- PROFIenergy energy-saving mode active'; 8802 'A08802 - PROFIenergy not possible to switch off incremental encoder supply'; 13009 'F13009 - Licensing OA application not licensed'; 13100 'F13100 - Know-how protection: Copy protection error'; 13101 'F13101 - Know-how protection: Copy protection cannot be activated'; 13102 'F13102 - Know-how protection: Consistency error of the protected data'; 30001 'F30001 - Power unit: Overcurrent'; 30002 'F30002 - Power unit: DC link voltage overvoltage'; 30003 'F30003 - Power unit: DC link voltage undervoltage'; 30004 'F30004 - Power unit: Overtemperature heat sink AC inverter'; 30005 'F30005 - Power unit: Overload I2t'; 30011 'F30011 - Power unit: Line phase failure in main circuit'; 30015 'F30015 (N, A) - Power unit: Phase failure motor cable'; 30016 'A30016 (N) - Power unit: Load supply switched out'; 30017 'F30017 - Power unit: Hardware current limit has responded too often'; 30021 'F30021 - Power unit: Ground fault'; 30022 'F30022 - Power unit: Monitoring U_ce'; 30024 'F30024 - Power unit: Overtemperature thermal model'; 30025 'F30025 - Power unit: Chip overtemperature'; 30027 'F30027 - Power unit: Precharging DC link time monitoring'; 30031 'A30031 - Power unit: Hardware current limiting in phase U'; 30032 'A30032 - Power unit: Hardware current limiting in phase V'; 30033 'A30033 - Power unit: Hardware current limiting in phase W'; 30034 'A30034 - Power unit: Internal overtemperature'; 30042 'A30042 - Power unit: Fan has reached the maximum operating hours'; 30051 'F30051 - Power unit: Motor holding brake short circuit detected'; 30052 'F30052 - EEPROM data error'; 30054 'A30054 (F, N) - Power unit: Undervoltage when opening the brake'; 30057 'A30057 - Power unit: Line asymmetry'; 30065 'A30065 (F, N) - Voltage measured values not plausible'; 30071 'F30071 - No new actual values received from the Power Module'; 30072 'F30072 - Setpoints can no longer be transferred to the Power Module'; 30074 'F30074 (A) - Communication error between the Control Unit and Power Module'; 30075 'F30075 - Configuration of the power unit unsuccessful'; 30080 'F30080 - Power unit: Current increasing too quickly'; 30081 'F30081 - Power unit: Switching operations too frequent'; 30105 'F30105 - PU: Actual value sensing fault'; 30502 'A30502 - Power unit: DC link overvoltage'; 30600 'F30600 - SI P2: STOP A initiated'; 30611 'F30611 (A) - SI P2: Defect in a monitoring channel'; 30620 'N30620 (F, A) - SI P2: Safe Torque Off active'; 30625 'F30625 - SI P2: Sign-of-life error in safety data'; 30649 'F30649 - SI P2: Internal software error'; 30650 'F30650 - SI P2: Acceptance test required'; 30651 'F30651 - SI P2: Synchronization with Control Unit unsuccessful'; 30655 'F30655 - SI P2: Align monitoring functions'; 30656 'F30656 - SI P2: Parameter processor 2 parameter error'; 30659 'F30659 - SI P2: Write request for parameter rejected'; 30662 'F30662 - Error in internal communications'; 30664 'F30664 - Error while booting'; 30665 'F30665 - SI P2: System is defective'; 30666 'A30666 (F) - SI Motion P2: Steady-state (static) 1 signal at the F-DI for safe acknowledgment'; 30680 'F30680 - SI Motion P2: Checksum error safety monitoring functions'; 30681 'F30681 - SI Motion P1: Incorrect parameter value'; 30682 'F30682 - SI Motion P2: Monitoring function not supported'; 30683 'F30683 - SI Motion P2: SLS enable missing'; 30692 'F30692 - SI Motion P2: Parameter value not permitted for encoderless'; 30693 'A30693 (F) - SI P2: Safety parameter settings changed, POWER ON required'; 30700 'C30700 - SI Motion P2: STOP A initiated'; 30701 'C30701 - SI Motion P2: STOP B initiated'; 30706 'C30706 - SI Motion P2: SAM/SBR limit exceeded'; 30711 'C30711 - SI Motion P2: Defect in a monitoring channel'; 30712 'C30712 - SI Motion P2: Defect in F-IO processing'; 30714 'C30714 - SI Motion P2: Safely limited speed exceeded'; 30716 'C30716 - SI Motion P2: Tolerance for safe motion direction exceeded'; 30770 'C30770 - SI Motion P2: Discrepancy error affecting the failsafe inputs'; 30772 'A30772 - SI Motion P2: Test stop for fail-safe digital outputs running'; 30773 'F30773 - SI Motion P2: Test stop fail-safe digital output error'; 30788 'A30788 - Automatic test stop: wait for STO deselection via SMM'; 30798 'C30798 - SI Motion P2: Test stop for motion monitoring functions running'; 30799 'C30799 - SI Motion P2: Acceptance test mode active'; 30800 'N30800 (F) - Power unit: Group signal'; 30802 'F30802 - Power unit: Time slice overflow'; 30804 'F30804 (N, A) - Power unit: CRC'; 30805 'F30805 - Power unit: EEPROM checksum error'; 30809 'F30809 - Power unit: Switching information not valid'; 30810 'A30810 (F) - Power unit: Watchdog timer'; 30850 'F30850 - Power unit: Internal software error'; 30903 'F30903 - Power unit: I2C bus error occurred'; 30920 'A30920 (F) - Temperature sensor fault'; 30950 'F30950 - Power unit: Internal software error'; 30999 'A30999 (F, N) - Power unit: Unknown alarm'; 31100 'F31100 (N, A) - Encoder 1: Zero mark distance error'; 31101 'F31101 (N, A) - Encoder 1: Zero mark failed'; 31103 'F31103 (N, A) - Encoder 1: Amplitude error track R'; 31118 'F31118 (N, A) - Encoder 1: Speed difference outside the tolerance range'; 31131 'F31131 (N, A) - Encoder 1: Deviation position incremental/absolute too large'; 31150 'F31150 (N, A) - Encoder 1: Initialization error'; 31153 'F31153 (N, A) - Encoder 1: Identification error'; 31400 'A31400 (F, N) - Encoder 1: Alarm threshold zero mark distance error'; 31401 'A31401 (F, N) - Encoder 1: Alarm threshold zero mark failed'; 31418 'A31418 (F, N) - Encoder 1: Speed difference per sampling rate exceeded'; 31422 'A31422 (F, N) - Encoder 1: Pulses per revolution square-wave encoder outside tolerance bandwidth'; 31431 'A31431 (F, N) - Encoder 1: Deviation position incremental/absolute too large'; 31802 'F31802 (N, A) - Encoder 1: Time slice overflow'; 31805 'F31805 (N, A) - Encoder 1: EEPROM checksum error'; 31850 'F31850 (N, A) - Encoder 1: Encoder evaluation internal software error'; 31899 'F31899 (N, A) - Encoder 1: Unknown fault'; 31905 'F31905 (N, A) - Encoder 1: Parameterization error'; 31915 'A31915 (F, N) - Encoder 1: Configuration error'; 31930 'A31930 (N) - Encoder 1: Data logger has saved data'; 31950 'F31950 - Encoder 1: Internal software error'; 31999 'A31999 (F, N) - Encoder 1: Unknown alarm'; 32110 'F32110 (N, A) - Encoder 2: Serial communications error'; 32111 'F32111 (N, A) - Encoder 2: Absolute encoder internal fault'; 32112 'F32112 (N, A) - Encoder 2: Error bit set in the serial protocol'; 32150 'F32150 (N, A) - Encoder 2: Initialization error'; 32153 'F32153 (N, A) - Encoder 2: Identification error'; 32410 'A32410 (F, N) - Encoder 2: Serial communications'; 32411 'A32411 (F, N) - Encoder 2: Absolute encoder signals internal alarms'; 32412 'A32412 (F, N) - Encoder 2: Error bit set in the serial protocol'; 32442 'A32442 (F, N) - Encoder 2: Battery voltage pre-alarm'; 32802 'F32802 (N, A) - Encoder 2: Time slice overflow'; 32805 'F32805 (N, A) - Encoder 2: EEPROM checksum error'; 32850 'F32850 (N, A) - Encoder 2: Encoder evaluation internal software error'; 32899 'F32899 (N, A) - Encoder 2: Unknown fault'; 32905 'F32905 (N, A) - Encoder 2: Parameterization error'; 32915 'A32915 (F, N) - Encoder 2: Configuration error'; 32930 'A32930 (N) - Encoder 2: Data logger has saved data'; 32950 'F32950 - Encoder 2: Internal software error'; 32999 'A32999 (F, N) - Encoder 2: Unknown alarm'; 50001 'A50001 (F) - PROFINET configuration error'; 50010 'A50010 (F) - PROFINET: Consistency error affecting adjustable parameters'; 50011 'A50011 (F) - Ethernet/IP: configuration error'; 50020 'A50020 (F) - PROFINET: Second controller missing'; 50510 'F50510 - FBLOCKS: Logon of the run-time group rejected'; 50511 'F50511 - FBLOCKS: Memory no longer available for free function blocks'; 50513 'A50513 (F) - FBLOCKS: Run sequence value already assigned'; 50517 'A50517 - FBLOCKS: Int. meas. active'; 50518 'F50518 - FBLOCKS: Sampling time of free run-time group differs at download'

text list "SDC_FAULTS-Old": 11 'Carrier 1 PLC Not Communicating'; 12 'Carrier 2 PLC Not Communicating'; 13 'Carrier 3 PLC Not Communicating'; 14 'Carrier 4 PLC Not Communicating'; 21 'Carrier 1 Safe Input Card Fault'; 22 'Carrier 1 Safe Output Card Fault'; 23 'Carrier 1 Standard Input Card Fault'; 24 'Carrier 1 Standard Output Card Fault'; 25 'Carrier 2 Safe Input Card Fault'; 26 'Carrier 2 Safe Output Card Fault'; 27 'Carrier 2 Standard Input Card Fault'; 28 'Carrier 2 Standard Output Card Fault'; 29 'Carrier 3 Safe Input Card Fault'; 30 'Carrier 3 Safe Output Card Fault'; 31 'Carrier 3 Standard Input Card Fault'; 32 'Carrier 3 Standard Output Card Fault'; 33 'Carrier 4 Safe Input Card Fault'; 34 'Carrier 4 Safe Output Card Fault'; 35 'Carrier 4 Standard Input Card Fault'; 36 'Carrier 4 Standard Output Card Fault'; 51 'Carrier 1 VFD Drive Fault'; 52 'Carrier 2 VFD Drive Fault'; 53 'Carrier 3 VFD Drive Fault'; 54 'Carrier 4 VFD Drive Fault'; 502 'Carrier 2 Crash Detection Fault'; 201 'Carrier 1 Encoder Reader Tilted 180 Degrees'; 202 'Carrier 1 Encoder Position Error'; 203 'Carrier 1 Encoder Internal Fault'; 211 'Carrier 2 Encoder Reader Tilted 180 Degrees'; 212 'Carrier 2 Encoder Position Error'; 213 'Carrier 2 Encoder Internal Fault'; 221 'Carrier 3 Encoder Reader Tilted 180 Degrees'; 222 'Carrier 3 Encoder Position Error'; 223 'Carrier 3 Encoder Internal Fault'; 231 'Carrier 4 Encoder Reader Tilted 180 Degrees'; 232 'Carrier 4 Encoder Position Error'; 233 'Carrier 4 Encoder Internal Fault'; 101 'Carrier 1 CB2120 Tripped'; 102 'Carrier 1 CB2121 Tripped'; 103 'Carrier 1 CB2122 Tripped'; 104 'Carrier 1 CB2123 Tripped'; 131 'Carrier 4 CB2120 Tripped'; 132 'Carrier 4 CB2121 Tripped'; 133 'Carrier 4 CB2122 Tripped'; 134 'Carrier 4 CB2123 Tripped'; 111 'Carrier 2 CB2120 Tripped'; 112 'Carrier 2 CB2121 Tripped'; 113 'Carrier 2 CB2122 Tripped'; 114 'Carrier 2 CB2123 Tripped'; 121 'Carrier 3 CB2120 Tripped'; 122 'Carrier 3 CB2121 Tripped'; 123 'Carrier 3 CB2122 Tripped'; 124 'Carrier 3 CB2123 Tripped'

text list "SDC_FAULTS": 24 'Scalance Ethernet SW2 Comm Fault'; 100 'Carrier 1 Profinet Comms Fault'; 101 'Carrier 1 Disconnect Open Power Fault DI11.0'; 102 'Carrier 1 CB02120 Tripped'; 103 'Carrier 1 CB02121 Tripped'; 104 'Carrier 1 CB02122 Tripped'; 105 'Carrier 1 CB02123 Tripped'; 106 'Carrier 1 AUX1 CB Tripped DI11.4'; 107 'Carrier 1 AUX2 CB Tripped DI11.5'; 111 'Carrier 1 PLC Not Communicating'; 121 'Carrier 1 Safe Input Card Fault'; 122 'Carrier 1 Safe Output Card Fault'; 123 'Carrier 1 Standard Input Card Fault'; 124 'Carrier 1 Standard Output Card Fault'; 130 'Carrier 1 PF Reader Tilted 180°'; 131 'Carrier 1 PF Reader Internal Error'; 132 'Carrier 1 PF Reader Position Error'; 133 'Carrier 1 PF Reader Comm Fault'; 134 'Carrier 1 FR HMI Comm Fault'; 140 'Carrier 1 Crash Detection Fault'; 145 'Carrier 1 Carrier Number Invalid'; 150 'F01653 - Carrier 1 SI P1 (CU): PROFIBUS/PROFINET configuration error'; 151 'F01662 - Carrier 1 Error internal communications'; 160 'F07011 - Carrier 1 Drive: Motor overtemperature'; 161 'F07016 - Carrier 1 Drive: Motor temperature sensor fault'; 162 'F07801 - Carrier 1 Drive: Motor overcurrent'; 163 'F07802 - Carrier 1 Drive: Infeed or power unit not ready'; 164 'F07807 - Carrier 1 Drive: Short-circuit/ground fault detected'; 170 'F08501 - Carrier 1 PROFINET: Setpoint timeout'; 180 'F30001 - Carrier 1 Power unit: Overcurrent'; 181 'F30002 - Carrier 1 Power unit: DC link voltage overvoltage'; 182 'F30003 - Carrier 1 Power unit: DC link voltage undervoltage'; 183 'F30004 - Carrier 1 Power unit: Overtemperature heat sink AC inverter'; 184 'F30005 - Carrier 1 Power unit: Overload I2t'; 185 'F30011 - Carrier 1 Power unit: Line phase failure in main circuit'; 186 'F30015 - Carrier 1 Power unit: Phase failure motor cable'; 20 'Rockwell PLC Comm Fault'; 21 'WLAN1 Comm Fault'; 22 'WLAN2 Comm Fault'; 23 'Scalance Ethernet SW1 Comm Fault'; 187 'F30021 - Carrier 1 Power unit: Ground fault'; 188 'F30024 - Carrier 1 Power unit: Overtemperature thermal model'; 189 'F30051 - Carrier 1 Power unit: Motor holding brake short circuit detected'; 200 'Carrier 2 Profinet Comms Fault'; 201 'Carrier 2 Disconnect Open Power Fault DI11.0'; 202 'Carrier 2 CB02120 Tripped'; 203 'Carrier 2 CB02121 Tripped'; 204 'Carrier 2 CB02122 Tripped'; 205 'Carrier 2 CB02123 Tripped'; 206 'Carrier 2 AUX1 CB Tripped DI11.4'; 207 'Carrier 2 AUX2 CB Tripped DI11.5'; 211 'Carrier 2 PLC Not Communicating'; 221 'Carrier 2 Safe Input Card Fault'; 222 'Carrier 2 Safe Output Card Fault'; 223 'Carrier 2 Standard Input Card Fault'; 224 'Carrier 2 Standard Output Card Fault'; 230 'Carrier 2 PF Reader Tilted 180°'; 231 'Carrier 2 PF Reader Position Error'; 232 'Carrier 2 PF Reader Internal Error'; 233 'Carrier 2 PF Reader Comm Fault'; 234 'Carrier 2 FR HMI Comm Fault'; 240 'Carrier 2 Crash Detection Fault'; 245 'Carrier 2 Carrier Number Invalid'; 250 'F01653 - Carrier 2 SI P1 (CU): PROFIBUS/PROFINET configuration error'; 251 'F01662 - Carrier 2 Error internal communications'; 260 'F07011 - Carrier 2 Drive: Motor overtemperature'; 261 'F07016 - Carrier 2 Drive: Motor temperature sensor fault'; 262 'F07801 - Carrier 2 Drive: Motor overcurrent'; 263 'F07802 - Carrier 2 Drive: Infeed or power unit not ready'; 264 'F07807 - Carrier 2 Drive: Short-circuit/ground fault detected'; 270 'F08501 - Carrier 2 PROFINET: Setpoint timeout'; 280 'F30001 - Carrier 2 Power unit: Overcurrent'; 281 'F30002 - Carrier 2 Power unit: DC link voltage overvoltage'; 282 'F30003 - Carrier 2 Power unit: DC link voltage undervoltage'; 283 'F30004 - Carrier 2 Power unit: Overtemperature heat sink AC inverter'; 284 'F30005 - Carrier 2 Power unit: Overload I2t'; 285 'F30011 - Carrier 2 Power unit: Line phase failure in main circuit'; 286 'F30015 - Carrier 2 Power unit: Phase failure motor cable'; 287 'F30021 - Carrier 2 Power unit: Ground fault'; 288 'F30024 - Carrier 2 Power unit: Overtemperature thermal model'; 289 'F30051 - Carrier 2 Power unit: Motor holding brake short circuit detected'; 300 'Carrier 3 Profinet Comms Fault'; 301 'Carrier 3 Disconnect Open Power Fault DI11.0'; 302 'Carrier 3 CB02120 Tripped'; 303 'Carrier 3 CB02121 Tripped'; 304 'Carrier 3 CB02122 Tripped'; 305 'Carrier 3 CB02123 Tripped'; 306 'Carrier 3 AUX1 CB Tripped DI11.4'; 307 'Carrier 3 AUX2 CB Tripped DI11.5'; 311 'Carrier 3 PLC Not Communicating'; 321 'Carrier 3 Safe Input Card Fault'; 322 'Carrier 3 Safe Output Card Fault'; 323 'Carrier 3 Standard Input Card Fault'; 324 'Carrier 3 Standard Output Card Fault'; 330 'Carrier 3 PF Reader Tilted 180°'; 331 'Carrier 3 PF Reader Position Error'; 332 'Carrier 3 PF Reader Internal Error'; 333 'Carrier 3 PF Reader Comm Fault'; 334 'Carrier 3 FR HMI Comm Fault'; 340 'Carrier 3 Crash Detection Fault'; 345 'Carrier 3 Carrier Number Invalid'; 350 'F01653 - Carrier 3 SI P1 (CU): PROFIBUS/PROFINET configuration error'; 351 'F01662 - Carrier 3 Error internal communications'; 360 'F07011 - Carrier 3 Drive: Motor overtemperature'; 361 'F07016 - Carrier 3 Drive: Motor temperature sensor fault'; 362 'F07801 - Carrier 3 Drive: Motor overcurrent'; 363 'F07802 - Carrier 3 Drive: Infeed or power unit not ready'; 364 'F07807 - Carrier 3 Drive: Short-circuit/ground fault detected'; 370 'F08501 - Carrier 3 PROFINET: Setpoint timeout'; 380 'F30001 - Carrier 3 Power unit: Overcurrent'; 381 'F30002 - Carrier 3 Power unit: DC link voltage overvoltage'; 382 'F30003 - Carrier 3 Power unit: DC link voltage undervoltage'; 383 'F30004 - Carrier 3 Power unit: Overtemperature heat sink AC inverter'; 384 'F30005 - Carrier 3 Power unit: Overload I2t'; 385 'F30011 - Carrier 3 Power unit: Line phase failure in main circuit'; 386 'F30015 - Carrier 3 Power unit: Phase failure motor cable'; 387 'F30021 - Carrier 3 Power unit: Ground fault'; 388 'F30024 - Carrier 3 Power unit: Overtemperature thermal model'; 389 'F30051 - Carrier 3 Power unit: Motor holding brake short circuit detected'; 400 'Carrier 4 Profinet Comms Fault'; 401 'Carrier 4 Disconnect Open Power Fault DI11.0'; 402 'Carrier 4 CB02120 Tripped'; 403 'Carrier 4 CB02121 Tripped'; 404 'Carrier 4 CB02122 Tripped'; 405 'Carrier 4 CB02123 Tripped'; 406 'Carrier 4 AUX1 CB Tripped DI11.4'; 407 'Carrier 4 AUX2 CB Tripped DI11.5'; 411 'Carrier 4 PLC Not Communicating'; 421 'Carrier 4 Safe Input Card Fault'; 422 'Carrier 4 Safe Output Card Fault'; 423 'Carrier 4 Standard Input Card Fault'; 424 'Carrier 4 Standard Output Card Fault'; 430 'Carrier 4 PF Reader Tilted 180°'; 431 'Carrier 4 PF Reader Position Error'; 432 'Carrier 4 PF Reader Internal Error'; 433 'Carrier 4 PF Reader Comm Fault'; 434 'Carrier 4 FR HMI Comm Fault'; 440 'Carrier 4 Crash Detection Fault'; 445 'Carrier 4 Carrier Number Invalid'; 450 'F01653 - Carrier 4 SI P1 (CU): PROFIBUS/PROFINET configuration error'; 451 'F01662 - Carrier 4 Error internal communications'; 460 'F07011 - Carrier 4 Drive: Motor overtemperature'; 461 'F07016 - Carrier 4 Drive: Motor temperature sensor fault'; 462 'F07801 - Carrier 4 Drive: Motor overcurrent'; 463 'F07802 - Carrier 4 Drive: Infeed or power unit not ready'; 464 'F07807 - Carrier 4 Drive: Short-circuit/ground fault detected'; 470 'F08501 - Carrier 4 PROFINET: Setpoint timeout'; 480 'F30001 - Carrier 4 Power unit: Overcurrent'; 481 'F30002 - Carrier 4 Power unit: DC link voltage overvoltage'; 482 'F30003 - Carrier 4 Power unit: DC link voltage undervoltage'; 483 'F30004 - Carrier 4 Power unit: Overtemperature heat sink AC inverter'; 484 'F30005 - Carrier 4 Power unit: Overload I2t'; 485 'F30011 - Carrier 4 Power unit: Line phase failure in main circuit'; 486 'F30015 - Carrier 4 Power unit: Phase failure motor cable'; 487 'F30021 - Carrier 4 Power unit: Ground fault'; 488 'F30024 - Carrier 4 Power unit: Overtemperature thermal model'; 489 'F30051 - Carrier 4 Power unit: Motor holding brake short circuit detected'; 10 'Carrier Spacing Fault'

graphic list "Grafikliste_G_Y": 0 'Green pilot light 2'; 1 'Yellow pilot light 2'

graphic list "PB_Slave_Bit12_3": 0 'PB_Array_blau_3'; 1 'PB_Array_grün_3'

graphic list "PB_Slave_Bit10_3": 0 'PB_Array_blau_3'; 1 'PB_Array_grün_3'

graphic list "PB_Slave_Bit7_3": 0 'PB_Array_blau_3'; 1 'PB_Array_grün_3'

graphic list "PB_Slave_Bit6_3": 1 'PB_Array_grün_3'; 0 'PB_Array_blau_3'

graphic list "PB_Slave_Bit5_3": 0 'PB_Array_blau_3'; 1 'PB_Array_grün_3'

graphic list "PB_Slave_Bit1_3": 1 'PB_Array_grün_3'; 0 'PB_Array_blau_3'

graphic list "PB_Slave_Bit3_3": 1 'PB_Array_grün_3'; 0 'PB_Array_blau_3'

graphic list "PB_Slave_Bit9_3": 0 'PB_Array_blau_3'; 1 'PB_Array_grün_3'

graphic list "PB_Slave_Bit8_3": 1 'PB_Array_grün_3'; 0 'PB_Array_blau_3'

graphic list "PB_Slave_Bit0_3": 1 'PB_Array_grün_3'; 0 'PB_Array_blau_3'

graphic list "PB_Slave_Bit4_3": 1 'PB_Array_grün_3'; 0 'PB_Array_blau_3'

graphic list "PB_Slave_Bit14_3": 0 'PB_Array_blau_3'; 1 'PB_Array_grün_3'

graphic list "PB_Slave_Bit11_3": 0 'PB_Array_blau_3'; 1 'PB_Array_grün_3'

graphic list "PB_Slave_Bit2_3": 1 'PB_Array_grün_3'; 0 'PB_Array_blau_3'

graphic list "PB_Slave_Bit13_3": 0 'PB_Array_blau_3'; 1 'PB_Array_grün_3'

graphic list "PB_Slave_Bit15_3": 1 'PB_Array_grün_3'; 0 'PB_Array_blau_3'

graphic list "PB_Slave_Bit1_1": 1 'PB_Array_grün_1'; 0 'PB_Array_blau_1'

graphic list "PB_Slave_Bit0_1": 1 'PB_Array_grün_1'; 0 'PB_Array_blau_1'

graphic list "PB_Slave_Bit2_1": 1 'PB_Array_grün_1'; 0 'PB_Array_blau_1'

graphic list "PB_Slave_Bit4_1": 1 'PB_Array_grün_1'; 0 'PB_Array_blau_1'

graphic list "PB_Slave_Bit3_1": 1 'PB_Array_grün_1'; 0 'PB_Array_blau_1'

graphic list "PB_Slave_Bit5_1": 0 'PB_Array_blau_1'; 1 'PB_Array_grün_1'

graphic list "PB_Slave_Bit7_1": 0 'PB_Array_blau_1'; 1 'PB_Array_grün_1'

graphic list "PB_Slave_Bit6_1": 1 'PB_Array_grün_1'; 0 'PB_Array_blau_1'

graphic list "PB_Slave_Bit13_1": 0 'PB_Array_blau_1'; 1 'PB_Array_grün_1'

graphic list "PB_Slave_Bit10_1": 0 'PB_Array_blau_1'; 1 'PB_Array_grün_1'

graphic list "PB_Slave_Bit12_1": 0 'PB_Array_blau_1'; 1 'PB_Array_grün_1'

graphic list "PB_Slave_Bit15_1": 1 'PB_Array_grün_1'; 0 'PB_Array_blau_1'

graphic list "PB_Slave_Bit9_1": 0 'PB_Array_blau_1'; 1 'PB_Array_grün_1'

graphic list "PB_Slave_Bit8_1": 1 'PB_Array_grün_1'; 0 'PB_Array_blau_1'

graphic list "PB_Slave_Bit11_1": 0 'PB_Array_blau_1'; 1 'PB_Array_grün_1'

graphic list "PB_Slave_Bit14_1": 0 'PB_Array_blau_1'; 1 'PB_Array_grün_1'

graphic list "PB_Slave_Bit4_2": 1 'PB_Array_grün_2'; 0 'PB_Array_blau_2'

graphic list "PB_Slave_Bit5_2": 0 'PB_Array_blau_2'; 1 'PB_Array_grün_2'

graphic list "PB_Slave_Bit7_2": 0 'PB_Array_blau_2'; 1 'PB_Array_grün_2'

graphic list "PB_Slave_Bit6_2": 1 'PB_Array_grün_2'; 0 'PB_Array_blau_2'

graphic list "PB_Slave_Bit2_2": 1 'PB_Array_grün_2'; 0 'PB_Array_blau_2'

graphic list "PB_Slave_Bit3_2": 1 'PB_Array_grün_2'; 0 'PB_Array_blau_2'

graphic list "PB_Slave_Bit1_2": 1 'PB_Array_grün_2'; 0 'PB_Array_blau_2'

graphic list "PB_Slave_Bit0_2": 1 'PB_Array_grün_2'; 0 'PB_Array_blau_2'

graphic list "PB_Slave_Bit14_2": 0 'PB_Array_blau_2'; 1 'PB_Array_grün_2'

graphic list "PB_Slave_Bit12_2": 0 'PB_Array_blau_2'; 1 'PB_Array_grün_2'

graphic list "PB_Slave_Bit15_2": 1 'PB_Array_grün_2'; 0 'PB_Array_blau_2'

graphic list "PB_Slave_Bit13_2": 0 'PB_Array_blau_2'; 1 'PB_Array_grün_2'

graphic list "PB_Slave_Bit10_2": 0 'PB_Array_blau_2'; 1 'PB_Array_grün_2'

graphic list "PB_Slave_Bit9_2": 0 'PB_Array_blau_2'; 1 'PB_Array_grün_2'

graphic list "PB_Slave_Bit8_2": 1 'PB_Array_grün_2'; 0 'PB_Array_blau_2'

graphic list "PB_Slave_Bit11_2": 0 'PB_Array_blau_2'; 1 'PB_Array_grün_2'

graphic list "@DiagnosticsStates": 0 '@Diagnostics_StateGood'; 1 '@Diagnostics_StateBad'

recipe "PN_100": Ort <- "PN_PB\Teiln_Nr_Ort", Typ <- "PN_PB\Teiln_Nr_Typ", Bezeichnung <- "PN_PB\Teiln_Nr_Bez"

recipe "PN_101": Ort <- "PN_PB\Teiln_Nr_Ort", Typ <- "PN_PB\Teiln_Nr_Typ", Bezeichnung <- "PN_PB\Teiln_Nr_Bez"

